   (* check and set outputs *)
     IF #X < #trigger_Low THEN
         #LOW := TRUE;
         #Status := 111;
         IF #Alarm_low THEN
             #Alarm := TRUE;
             #Status := 1;
         END_IF;
     ELSIF #X < #T_1 THEN
         #Q1 := TRUE;
     ELSIF #X < #T_2 THEN
         #Q2 := TRUE;
     ELSIF #X < #T_3 THEN
         #Q3 := TRUE;
     ELSIF #X < #T_4 THEN
         #Q4 := TRUE;
     ELSIF #X < #T_5 THEN
         #Q5 := TRUE;
     ELSIF #X < #trigger_High THEN
         #Q6 := TRUE;
     ELSE
         #HIGH := TRUE;
         #Status := 112;
         IF #Alarm_high THEN
             #Alarm := TRUE;
             #Status := 2;
         END_IF;
     END_IF;

   (* revision history
   hm  22. feb 2007  rev 1.0
     original version

   hm  2. dec 2007   rev 1.1
     chaged code for better performance

   hm  6. jan 2008   rev 1.2
     further performance improvement

   *)
END_FUNCTION_BLOCK

FUNCTION_BLOCK "CALIBRATE"   // FB124, SCL
TITLE = CALIBRATE
{ S7_Optimized_Access := 'FALSE' }
AUTHOR : hugo
FAMILY : MEASURE
NAME : CALIBR
VERSION : 1.3
// Calibrate allows for offset and scale calibration of an analog input.
// offset is calibrated to a stored reference Y_offset while CO is true.
// after the offset is calibrated, scale can be calibrated to a reference value Y_scale while CS is true.
   VAR_INPUT
      X : Real;
      CO : Bool;
      CS : Bool;
      Y_Offset : Real;
      Y_Scale : Real;
   END_VAR
   VAR_OUTPUT
      Y : Real;
   END_VAR
   VAR
      offset : Real;
      Scale : Real := 1.0e+0;
   END_VAR
BEGIN


   (* check for calibration *)
   IF #CO THEN
       #offset := #Y_Offset - #X;
   ELSIF #CS THEN
       #Scale := #Y_Scale / (#X + #offset);
   END_IF;
   (* calculate output *)
   #Y := (#X + #offset) * #Scale;


   (* revision history
   hm 22.2.2007        rev 1.2
       changed VAR RETAIN PERSISTENT to VAR RETAIN for better compatibility
       wago lon contollers do not support persisitent

   hm  11. mar. 2009   rev 1.3
       changed real constants to use dot syntax

   *)
END_FUNCTION_BLOCK

FUNCTION_BLOCK "CYCLE_TIME"   // FB125, SCL
TITLE = CYCLE_TIME
{ S7_Optimized_Access := 'FALSE' }
AUTHOR : hugo
FAMILY : MEASURE
NAME : CYCLE
VERSION : 1.2
// this function block measures the cycle time and displays the last, min and max cycle time of the current task.
// the resolution is 1ms.
// the cycles output is a dword counter which counts the cycles.
// a rst pulse on the input will reset all data.
// 
// uses: T_PLC_MS [FC64]
//       STIME [FB64],IDB_STIME [DB64]
   VAR_INPUT
      rst : Bool;
   END_VAR
   VAR_OUTPUT
      ct_min : Time;
      ct_max : Time;
      ct_last : Time;
      systime : Time;
      sysdays : Int;
      cycles : DWord;
   END_VAR
   VAR
      last_cycle : Time;
      tx : Time;
      init : Bool;
   END_VAR
   VAR_TEMP
      TOP_SI : Struct
         EV_CLASS : Byte;
         EV_NUM : Byte;
         PRIORITY : Byte;
         NUM : Byte;
         TYP2_3 : Byte;
         TYP1 : Byte;
         ZI1 : Word;
         ZI2_3 : DWord;
      END_STRUCT;
      START_UP_SI : Struct
         EV_CLASS : Byte;
         EV_NUM : Byte;
         PRIORITY : Byte;
         NUM : Byte;
         TYP2_3 : Byte;
         TYP1 : Byte;
         ZI1 : Word;
         ZI2_3 : DWord;
      END_STRUCT;
      ERR : Int;
   END_VAR
BEGIN


   (* read actual startup info *)
   (* OB1_SCAN_1  BYTE  -  B#16#01: Abschluss des Neustarts (Warmstarts)
                        -  B#16#02: Abschluss des Wiederanlaufs
                        -  B#16#03: Abschluss des freien Zyklus
                        -  B#16#04: Abschluss des Kaltstarts
                        -  B#16#05: Erster OB 1-Zyklus der neuen Master-CPU nach 
                                    Master-Reserve-Umschaltung und STOP des 
                                    bisherigen Masters *)

     #ERR := RD_SINFO (TOP_SI => #TOP_SI, START_UP_SI => #START_UP_SI);

   (* reset last_time on system startup *)
     IF #TOP_SI.EV_NUM <> 3 THEN 
       #last_cycle := t#0ms;
     END_IF;

     #tx := T_CONV(DWORD_TO_DINT("T_PLC_MS"())) - #last_cycle;

     IF #rst THEN
         #ct_min := t#10h;
         #ct_max := t#0ms;
         #cycles := 0;
     ELSIF #last_cycle > t#0s THEN
         IF #tx < #ct_min THEN #ct_min := #tx;
         ELSIF #tx > #ct_max THEN #ct_max := #tx;
         END_IF;
         #ct_last := #tx;
     ELSIF #ct_min = t#0s THEN
         #ct_min := t#0s - t#1ms;
     END_IF;
     IF #init THEN
         #systime := #systime + #tx;
             IF #systime >= t#1d THEN
                 #systime := #systime - t#1d;
                 #sysdays := #sysdays + 1;
             END_IF;
     END_IF;
     #init := TRUE;
     #last_cycle := #last_cycle + #tx;
     #cycles := DINT_TO_DWORD(DWORD_TO_DINT(#cycles) + 1);

   (*    revision history
   hm 12.12.2006        rev 1.1
       added cycles output, a dword cycle counter.
   hm 10.3.2007         rev 1.2
       changed initialization of ct_min to t#10h for compatibility with siemens s7

   *)
END_FUNCTION_BLOCK

FUNCTION_BLOCK "DT_SIMU"   // FB126, SCL
TITLE = DT_SIMU
{ S7_Optimized_Access := 'FALSE' }
AUTHOR : hugo
FAMILY : MEASURE
NAME : DTSIMU
VERSION : 1.2
// DT_SIMU simulates a real time clock and can be adjusted to different speeds
// it can also be used in simulation to simulate a real time clock.
// the peed of the clock can be increased or decreased to debug timers.
// with the input start a start date-time can be specified.
// 
// uses: AD_DT_TM [FC1]
//       T_PLC_MS [FC64]
//       STIME [FB64],IDB_STIME [DB64]
   VAR_INPUT
      START : Date_And_Time;
      SPEED : Real := 1.0e+0;
   END_VAR
   VAR_OUTPUT
      DTS : Date_And_Time;
   END_VAR
   VAR
      tc : DWord;
      init : Bool;
      last : DWord;
      tx : DWord;
      td : DWord;
   END_VAR
   VAR_TEMP
      TOP_SI : Struct
         EV_CLASS : Byte;
         EV_NUM : Byte;
         PRIORITY : Byte;
         NUM : Byte;
         TYP2_3 : Byte;
         TYP1 : Byte;
         ZI1 : Word;
         ZI2_3 : DWord;
      END_STRUCT;
      START_UP_SI : Struct
         EV_CLASS : Byte;
         EV_NUM : Byte;
         PRIORITY : Byte;
         NUM : Byte;
         TYP2_3 : Byte;
         TYP1 : Byte;
         ZI1 : Word;
         ZI2_3 : DWord;
      END_STRUCT;
      ERR : Int;
   END_VAR
BEGIN


   (* read actual startup info *)
   (* OB1_SCAN_1  BYTE  -  B#16#01: Abschluss des Neustarts (Warmstarts)
                        -  B#16#02: Abschluss des Wiederanlaufs
                        -  B#16#03: Abschluss des freien Zyklus
                        -  B#16#04: Abschluss des Kaltstarts
                        -  B#16#05: Erster OB 1-Zyklus der neuen Master-CPU nach 
                                    Master-Reserve-Umschaltung und STOP des 
                                    bisherigen Masters *)

   #ERR := RD_SINFO (TOP_SI => #TOP_SI, START_UP_SI => #START_UP_SI);

   (* reset last_time on system startup *)
   IF #TOP_SI.EV_NUM = 1 OR #TOP_SI.EV_NUM = 2 OR #TOP_SI.EV_NUM = 4 THEN 
       #init := FALSE;
   END_IF;

   (* read system timer *)
   #tx := "T_PLC_MS"();
   #tc := DINT_TO_DWORD(REAL_TO_DINT(DINT_TO_REAL((DWORD_TO_DINT(#tx) - DWORD_TO_DINT(#last))) * #SPEED));

   IF NOT #init THEN
       #init := TRUE;
       #DTS := #START;
       #tc := 0;
       #last := #tx;
   ELSIF #SPEED = 0.0 THEN
       #DTS := #DTS T_ADD T_CONV(1);
   ELSIF DWORD_TO_DINT(#tc) >= 1000 THEN
       #td := DINT_TO_DWORD((DWORD_TO_DINT(#tc) / 1000)*1000);
       #DTS := #DTS T_ADD T_CONV(DWORD_TO_DINT(#td));
       #last := DINT_TO_DWORD(DWORD_TO_DINT(#last) + REAL_TO_DINT(DINT_TO_REAL(DWORD_TO_DINT(#td)) / #SPEED));
   END_IF;


   (* revision history
   hm  11. sep. 2008   rev 1.0
       original version

   hm  16. nov 2008    rev 1.1
       added type conversions for compatibility reasons

   hm  8.  mar. 2009   rev 1.2
       added increment by cycle mode

   *)
END_FUNCTION_BLOCK

FUNCTION_BLOCK "METER"   // FB127, SCL
TITLE = METER
{ S7_Optimized_Access := 'FALSE' }
AUTHOR : oscat
FAMILY : MEASURE
NAME : METER
VERSION : 1.4
// METER measures usage of power or similar values the output MX is the sum of the inputs over time.
// MX := sum over time of (I1 * P1 + I2 * P2)/D.
// a simple example is the consumption counter for a 2 stage oil burner where stage 1 is 10KW and stage 2 is 20KW.
// I1 and I2 decide which value is accounted for, I1 = True only counts P1, I2 is True counts P2 
// and I1 and I2 is true counts P1 and P2.
// the meter can be used for all kind of consumption meters. P1 and P2 can change on the fly.
// 
// uses: REAL2 [UDT11]
//       T_PLC_MS [FC64]
//       STIME [FB64],IDB_STIME [DB64]
//       R2_ADD [FC144]
   VAR_INPUT
      M1 : Real;
      M2 : Real;
      I1 : Bool;
      I2 : Bool;
      D : Real := 1.0e+0;
      RST : Bool;
   END_VAR
   VAR_IN_OUT
      MX : Real;
   END_VAR
   VAR
      MR : "REAL2";
      MX1 : Real;
      MX2 : Real;
      tx : DWord;
      last : DWord;
      tc : Real;
      init : Bool;
   END_VAR
   VAR_TEMP
      TOP_SI : Struct
         EV_CLASS : Byte;
         EV_NUM : Byte;
         PRIORITY : Byte;
         NUM : Byte;
         TYP2_3 : Byte;
         TYP1 : Byte;
         ZI1 : Word;
         ZI2_3 : DWord;
      END_STRUCT;
      START_UP_SI : Struct
         EV_CLASS : Byte;
         EV_NUM : Byte;
         PRIORITY : Byte;
         NUM : Byte;
         TYP2_3 : Byte;
         TYP1 : Byte;
         ZI1 : Word;
         ZI2_3 : DWord;
      END_STRUCT;
      ERR : Int;
   END_VAR
BEGIN


   (* read actual startup info *)
   (* OB1_SCAN_1  BYTE  -  B#16#01: Abschluss des Neustarts (Warmstarts)
                        -  B#16#02: Abschluss des Wiederanlaufs
                        -  B#16#03: Abschluss des freien Zyklus
                        -  B#16#04: Abschluss des Kaltstarts
                        -  B#16#05: Erster OB 1-Zyklus der neuen Master-CPU nach 
                                    Master-Reserve-Umschaltung und STOP des 
                                    bisherigen Masters *)

   #ERR := RD_SINFO (TOP_SI => #TOP_SI, START_UP_SI => #START_UP_SI);

   (* reset last_time on system startup *)
   IF #TOP_SI.EV_NUM = 1 OR #TOP_SI.EV_NUM = 2 OR #TOP_SI.EV_NUM = 4 THEN 
       #init := FALSE;
   END_IF;

   (* measure the last cycle time and make sure we onle execute once every millisecond *)
   #tx := "T_PLC_MS"();

   IF NOT #init THEN
       #init := TRUE;
       #last := #tx;
       #MR.RX := #MX;
       #MR.R1 := 0.0;
   ELSIF #tx = #last THEN
       RETURN;
   ELSE
       #tc := DINT_TO_REAL(DWORD_TO_DINT(#tx) - DWORD_TO_DINT(#last)) * 0.001;
   END_IF;
   #last := #tx;

   (* reset *)
   IF #RST THEN
       #MR.R1 := 0.0;
       #MR.RX := 0.0;
   ELSE
       (* current consumption measurement *)
       IF #I1 THEN #MX1 := #M1; ELSE #MX1 := 0.0; END_IF;
       IF #I2 THEN #MX2 := #M2; ELSE #MX2 := 0.0; END_IF;
       (* add up the current values in a double real *)
       #MR := "R2_ADD"(X:=#MR,Y:=(SEL(G:=#I1,IN0:=0.0,IN1:=#MX1) + SEL(G:=#I2,IN0:=0.0,IN1:=#MX2)) / #D * #tc);
       (* set the current output value *)
       #MX := #MR.RX;
   END_IF;


   (* revision history

   hm  16. sep.2007        rev 1.0
       original version

   hm  7. feb 2008     rev 1.1
       use new version of ft_int to avoid a counting stop at high values
       deleted unnecessary limits

   hm  24. mar. 2008   rev 1.2
       use data_type real2 to extend accuracy to 15 digits total
       do not use ft_int which adds unnecessary overhead

   hm  8. feb. 2009    rev 1.3
       changed mx to be I/O
       make sure calculation works for cycle times < 1 ms

   hm  8. mar. 2009    rev 1.4
       last was not updated
       code improvements

   *)
END_FUNCTION_BLOCK

FUNCTION_BLOCK "METER_STAT"   // FB128, SCL
TITLE = METER_STAT
{ S7_Optimized_Access := 'FALSE' }
AUTHOR : oscat
FAMILY : MEASURE
NAME : METER_ST
VERSION : 1.3
// METER_STAT runs statistics of a metered value, it calculates the current week, day, month and year consumption and stores the corresponding last day, week, month and year value.
// 
// uses: YEAR_OF_DATE [FC219]
//       MONTH_OF_DATE [FC202]
//       DAY_OF_YEAR [FC180]
//       YEAR_BEGIN [FC217]
//       YEAR_OF_DATE [FC219]
//       LEAP_OF_DATE [FC193] 
//       LEAP_YEAR [FC194]
//       DAY_OF_WEEK [FC179]
   VAR_INPUT
      IN : Real;
      _DI : Date;
      RST : Bool;
   END_VAR
   VAR_IN_OUT
      Last_Day : Real;
      Current_Day : Real;
      Last_Week : Real;
      Current_Week : Real;
      Last_Month : Real;
      Current_Month : Real;
      Last_Year : Real;
      Current_Year : Real;
   END_VAR
   VAR
      Year_Start : Real;
      Month_Start : Real;
      Week_Start : Real;
      Day_Start : Real;
      last_run : Date;
   END_VAR
BEGIN


   IF #RST THEN
       #Last_Day := 0.0;
       #Current_Day := 0.0;
       #Day_Start := #IN;
       #Last_Week := 0.0;
       #Current_Week := 0.0;
       #Week_Start := #IN;
       #Last_Month := 0.0;
       #Current_Month := 0.0;
       #Month_Start := #IN;
       #Last_Year := 0.0;
       #Current_Year := 0.0;
       #Year_Start := #IN;
   ELSE
       #Current_Day := #IN - #Day_Start;
       #Current_Week := #IN - #Week_Start;
       #Current_Month := #IN - #Month_Start;
       #Current_Year := #IN - #Year_Start;
   END_IF;

   IF "YEAR_OF_DATE"(#_DI) > "YEAR_OF_DATE"(#last_run) THEN
       (* a new year has started *)
       #Last_Year := #Current_Year;
       #Current_Year := 0.0;
       #Year_Start := #IN;
       #Last_Month := #Current_Month;
       #Current_Month := 0.0;
       #Month_Start := #IN;
       #Last_Day := #Current_Day;
       #Current_Day := 0.0;
       #Day_Start := #IN;
   ELSIF "MONTH_OF_DATE"(#_DI) > "MONTH_OF_DATE"(#last_run) THEN
       (* a new month has started, january is alrerady done by year change *)
       #Last_Month := #Current_Month;
       #Current_Month := 0.0;
       #Month_Start := #IN;
       #Last_Day := #Current_Day;
       #Current_Day := 0.0;
       #Day_Start := #IN;
   ELSIF "DAY_OF_YEAR"(#_DI) > "DAY_OF_YEAR"(#last_run) THEN
       (* day has chaged, first day of year and first day of month has already been taken care of *)
       #Last_Day := #Current_Day;
       #Current_Day := 0.0;
       #Day_Start := #IN;
   END_IF;
   IF "DAY_OF_WEEK"(#_DI) < "DAY_OF_WEEK"(#last_run) THEN
       (* a new week has started *)
       #Last_Week := #Current_Week;
       #Current_Week := 0.0;
       #Week_Start := #IN;
   END_IF;
   #last_run := #_DI;


   (* revision history
   hm  16. sep. 2007 rev 1.0
     original version

   hm  7. oct. 2008  rev 1.1
     changed function year_to_year_of_date
     changed function month to month_of_date
     changed function weekday to day_of_week

   hm  11. mar. 2009 rev 1.2
     changed real constants to use dot syntax

   hm  18. jul. 2009 rev 1.3
     changes all outputs to be I/O
   *)
END_FUNCTION_BLOCK

FUNCTION_BLOCK "M_D"   // FB129, SCL
TITLE = M_D
{ S7_Optimized_Access := 'FALSE' }
AUTHOR : hugo
FAMILY : MEASURE
NAME : M_D
VERSION : 1.2
// m_d measures the time between a rising edge on start to a rising edge on stop and returs the last measured value on the output PT.
// a second output ET is starting from 0 at the rising edge of start and is counting up until the rising edge of stop occurs.
// the asynchronous input rst can reset the outputs at any time.
// tmax defines a timeout wich is the maximum measurable time between start and stop, if this time is exceeded the outputs will stay at 0.
// 
// uses: T_PLC_MS [FC64]
//       STIME [FB64],IDB_STIME [DB64]
   VAR_INPUT
      start : Bool;
      stop : Bool;
      tmax : Time := T#10D;
      rst : Bool;
   END_VAR
   VAR_OUTPUT
      PT : Time;
      ET : Time;
      run : Bool;
   END_VAR
   VAR
      edge : Bool;
      T_0 : Time;
      tx : Time;
      startup : Bool;
   END_VAR
   VAR_TEMP
      TOP_SI : Struct
         EV_CLASS : Byte;
         EV_NUM : Byte;
         PRIORITY : Byte;
         NUM : Byte;
         TYP2_3 : Byte;
         TYP1 : Byte;
         ZI1 : Word;
         ZI2_3 : DWord;
      END_STRUCT;
      START_UP_SI : Struct
         EV_CLASS : Byte;
         EV_NUM : Byte;
         PRIORITY : Byte;
         NUM : Byte;
         TYP2_3 : Byte;
         TYP1 : Byte;
         ZI1 : Word;
         ZI2_3 : DWord;
      END_STRUCT;
      ERR : Int;
   END_VAR
BEGIN


   (* read actual startup info *)
   (* OB1_SCAN_1  BYTE  -  B#16#01: Abschluss des Neustarts (Warmstarts)
                        -  B#16#02: Abschluss des Wiederanlaufs
                        -  B#16#03: Abschluss des freien Zyklus
                        -  B#16#04: Abschluss des Kaltstarts
                        -  B#16#05: Erster OB 1-Zyklus der neuen Master-CPU nach 
                                    Master-Reserve-Umschaltung und STOP des 
                                    bisherigen Masters *)

   #ERR := RD_SINFO (TOP_SI => #TOP_SI, START_UP_SI => #START_UP_SI);

   (* reset last_time on system startup *)
   IF #TOP_SI.EV_NUM <> 3 THEN 
       #T_0 := t#0ms;
   END_IF;

   (* check for rst input *)
   IF #rst OR #ET >= #tmax THEN
       #PT := t#0ms;
       #ET := t#0ms;
       #startup := FALSE;
       #run := FALSE;
   END_IF;

   (* avoid timers to start when input is true at startup *)
   IF NOT #startup THEN
       #edge := #start;
       #startup := TRUE;
   END_IF;

   (* read system timer *)
   #tx := T_CONV(DWORD_TO_DINT("T_PLC_MS"()));

   (* detect rising edge on start *)
   IF #start AND NOT #edge AND NOT #stop THEN
       #T_0 := #tx;
       #run := TRUE;
       #PT := t#0s;
   ELSIF #stop AND #run THEN
       #PT := #ET;
       #run := FALSE;
   END_IF;
   #edge := #start;
   IF #run THEN #ET := #tx - #T_0; END_IF;


   (* revision history
   hm      2.5.2007    rev 1.0
       original version

   hm        16.9.2007   rev 1.1
       changes time() to T_plc_ms() for compatibility reasons

   hm  27. feb 2009    rev 1.2
       deleted unnecessary init with 0
   *)
END_FUNCTION_BLOCK

FUNCTION_BLOCK "M_T"   // FB130, SCL
TITLE = M_T
{ S7_Optimized_Access := 'FALSE' }
AUTHOR : hugo
FAMILY : MEASURE
NAME : M_T
VERSION : 1.4
// m_t measures the with of a high pulse and returs the last measured pulse width on output PT.
// a second output ET is starting from 0 at the rising edge and counting up until the falling edge occurs and resetts et to 0.
// the asynchrtonous input rst can reset the outputs at any time.
// tmax defines a maximum measurable time, if this value is exceeded the outputs will be reset to 0.
// 
// uses: T_PLC_MS [FC64]
//       STIME [FB64],IDB_STIME [DB64]
   VAR_INPUT
      IN : Bool;
      TMAX : Time := T#10D;
      RST : Bool;
   END_VAR
   VAR_OUTPUT
      PT : Time;
      ET : Time;
   END_VAR
   VAR
      edge : Bool;
      start : Time;
      tx : Time;
   END_VAR
BEGIN


   #tx := T_CONV(DWORD_TO_DINT("T_PLC_MS"()));

   IF #RST OR #ET >= #TMAX THEN
       #PT := t#0s; 
       #ET := t#0s;
   ELSIF #IN THEN
       IF NOT #edge THEN #start := #tx; END_IF;
       #ET := #tx - #start;
   ELSE
       #PT := #ET;
   END_IF;
   #edge := #IN;


   (* revision history
   hm  4. aug. 2006    rev 1.0
       original version

   hm  2. may. 2007    rev 1.1
       added init variable to avoid unreasonable measurement if falling edge occurs first.
       added et (elapsed time) output to count from 0 at rising edge until a falling edge resets et to 0.
       added reset input.

   hm  16. sep. 2007   rev 1.2
       changes time() to T_plc_ms() for compatibility reasons

   hm  17. dec. 2008   rev 1.3
       code optimized

   hm  10. mar. 2009   rev 1.4
       removed nested comments
       removed double assignments

   *)
END_FUNCTION_BLOCK

FUNCTION_BLOCK "M_TX"   // FB131, SCL
TITLE = M_TX
{ S7_Optimized_Access := 'FALSE' }
AUTHOR : oscat
FAMILY : MEASURE
NAME : M_TX
VERSION : 1.4
// this measures the timing of a signal
// TH is the high pulse width
// TL is the low pulse width
// DC is the duty cycle
// F is the frequency
// ET will start at 0 with a rising edge and count up till the next rising edge starts from 0 again. 
// the acuracy depends on the cycle time of the sps and is limited to 1ms resolution.
// an asynchronous reset can reset all outputs to 0 at any time.
// the input tmax can configure a timeout for ET where the function block will outomatically reset itself.
// tmx is predefined to 10 days.
// 
// uses: T_PLC_MS [FC64]
//       STIME [FB64],IDB_STIME [DB64]
   VAR_INPUT
      in : Bool;
      tmax : Time := T#10D;
      rst : Bool;
   END_VAR
   VAR_OUTPUT
      TH : Time;
      TL : Time;
      DC : Real;
      F : Real;
      ET : Time;
   END_VAR
   VAR
      edge : Bool;
      start : Time;
      stop : Time;
      tx : Time;
      rise : Bool;
      fall : Bool;
      startup : Bool;
   END_VAR
BEGIN


   (* check FOR rst input *)
   IF #rst OR (#ET >= #tmax) THEN
       #rise := FALSE;
       #fall := FALSE;
       #startup := FALSE;
       #TH := t#0ms;
       #TL := t#0ms;
       #DC := 0.0;
       #F := 0.0;
       #ET := t#0s;
   END_IF;

   (* avoid timers to start when input is true at startup *)
   IF NOT #startup THEN
       #edge := #in;
       #startup := TRUE;
   END_IF;

   (* read system timer *)
   #tx := T_CONV(DWORD_TO_DINT("T_PLC_MS"()));

   (* edge trigger rising and falling edge *)
   IF #in XOR #edge THEN
       #edge := #in;
       (* rising edge starts measurement *)
       IF #in THEN
           #start := #tx;
           #rise := TRUE;
           IF #fall THEN #TL := #start - #stop; END_IF;
           IF #TH > t#0ms AND #TL > t#0ms THEN
               #DC := DINT_TO_REAL(T_CONV(#TH)) / DINT_TO_REAL(T_CONV(#TH+#TL));
               #F := 1000.0 / DINT_TO_REAL(T_CONV(#TH + #TL));
           END_IF;
       (* falling edge starts second cycle measurement *)
       ELSE
           #stop := #tx;
           #fall := TRUE;
           IF #rise THEN #TH := #stop - #start; END_IF;
           IF #TH > t#0ms AND #TL > t#0ms THEN
               #DC := DINT_TO_REAL(T_CONV(#TH)) /  DINT_TO_REAL(T_CONV(#TH+#TL));
               #F := 1000.0 / DINT_TO_REAL(T_CONV(#TH + #TL));
           END_IF;
       END_IF;
   END_IF;
   IF #rise THEN #ET := #tx - #start; END_IF;


   (* revision history
   hm  4. aug. 2006    rev 1.0
       original version

   hm  2. mai. 2007    rev 1.1
       made sure that no undefined values would be measured at startup conditions
       added output et
       added rst input
       added tmax input

   hm  16. sep. 2007   rev 1.2
       changes time() to T_plc_ms() for compatibility reasons

   hm  27. feb. 2009   rev 1.3
       deleted unnecessary init with 0

   hm  11. mar. 2009   rev 1.4
       changed real constants to use dot syntax

   *)
END_FUNCTION_BLOCK

FUNCTION_BLOCK "ONTIME"   // FB132, SCL
TITLE = ONTIME
{ S7_Optimized_Access := 'FALSE' }
AUTHOR : oscat
FAMILY : MEASURE
NAME : ONTIME
VERSION : 2.5
// ONTIME measures the ontime of a signal in seconds.
// the output SECONDS is of type DWORD which results in a total measurement range of 1 second up to 136 years.
// internally ontime works with a resolution of milliseconds
// 
// uses: T_PLC_MS [FC64]
//       STIME [FB64],IDB_STIME [DB64]
   VAR_INPUT
      IN : Bool;
      RST : Bool;
   END_VAR
   VAR_IN_OUT
      SECONDS : DInt;
      CYCLES : DInt;
   END_VAR
   VAR
      tx : DWord;
      last : DWord;
      edge : Bool;
      init : Bool;
      ms : DWord;
   END_VAR
   VAR_TEMP
      TOP_SI : Struct
         EV_CLASS : Byte;
         EV_NUM : Byte;
         PRIORITY : Byte;
         NUM : Byte;
         TYP2_3 : Byte;
         TYP1 : Byte;
         ZI1 : Word;
         ZI2_3 : DWord;
      END_STRUCT;
      START_UP_SI : Struct
         EV_CLASS : Byte;
         EV_NUM : Byte;
         PRIORITY : Byte;
         NUM : Byte;
         TYP2_3 : Byte;
         TYP1 : Byte;
         ZI1 : Word;
         ZI2_3 : DWord;
      END_STRUCT;
      ERR : Int;
   END_VAR
BEGIN


     (* read actual startup info *)
     (* OB1_SCAN_1  BYTE  -  B#16#01: Abschluss des Neustarts (Warmstarts)
                          -  B#16#02: Abschluss des Wiederanlaufs
                          -  B#16#03: Abschluss des freien Zyklus
                          -  B#16#04: Abschluss des Kaltstarts
                          -  B#16#05: Erster OB 1-Zyklus der neuen Master-CPU nach 
                                      Master-Reserve-Umschaltung und STOP des 
                                      bisherigen Masters *)

     #ERR := RD_SINFO (TOP_SI => #TOP_SI, START_UP_SI => #START_UP_SI);

     (* read system time *)
     #tx := "T_PLC_MS"();

     (* reset last_time on system startup *)
     IF #TOP_SI.EV_NUM = 1 OR #TOP_SI.EV_NUM = 2 OR #TOP_SI.EV_NUM = 4 THEN 
         #init := FALSE;
     END_IF;

     (* make sure the first cycle works correctly *)
     IF NOT #init THEN
       #init := TRUE;
       #last := #tx;
       #ms := 0;
     END_IF;
     IF #RST THEN
       #SECONDS := 0;
       #CYCLES := 0;
       #last := #tx;
       #ms := 0;
     ELSIF #IN THEN
       (* add the current milliseconds *)
       #ms := DINT_TO_DWORD((DWORD_TO_DINT(#tx) - DWORD_TO_DINT(#last)) + DWORD_TO_DINT(#ms));
       IF DWORD_TO_DINT(#ms) >= 1000 THEN
         #SECONDS := #SECONDS + 1;
         #ms := DINT_TO_DWORD(DWORD_TO_DINT(#ms) - 1000);
       END_IF;
       #CYCLES := #CYCLES + BOOL_TO_DINT(NOT #edge);
     END_IF;
     #last := #tx;
     #edge := #IN;


   (* revision history
   hm 22.2.2007    rev 1.1
     changed VAR RETAIN PERSISTENT to VAR RETAIN for better compatibility
     wago lon contollers do not support persisitent

   hm 2.8.2007   rev 1.2
     adding time up in a real number will automatically lead to the point where 
     small time scales like the cycle time will be below the resolution of real and therefore
     ontime would not increase in small steps as necessary
     the time is now measured internally in two  dwords and be converted to real only for
     output purposes.
     deleted the variable power because it was unnecessary

   hm  16.9.2007   rev 1.3
     changes time() to T_plc_ms() for compatibility reasons

   hm  2. dec. 2007  rev 1.4
     chaged code for better performance

   hm  16. mar. 2008 rev 1.5
     added type conversions to avoid warnings under codesys 3.0

   hm  21. oct. 2008 rev 2.0
     changed module for much better performance and allow for external result storage

   hm  10. nov. 2008 rev 2.1
     increased internal resolution to milliseconds

   hm  16. nov. 2008 rev 2.2
     changed typecast to avoid warnings

   hm  17. dec. 2008 rev 2.3
     fixed an error when in would be true for more then 49 days

   hm  17. jan 2011  rev 2.4
     init will not clear seconds and cycles, only rst clears these values  

   hm  18. mar. 2011 rev 2.5
     reset was not working

   *)
END_FUNCTION_BLOCK

FUNCTION_BLOCK "TC_MS"   // FB133, SCL
TITLE = TC_MS
{ S7_Optimized_Access := 'FALSE' }
AUTHOR : hugo
FAMILY : MEASURE
NAME : TC_MS
VERSION : 1.0
// TC_MS delivers the time it was last called on the output TC in Milliseconds.
// 
// uses: T_PLC_MS [FC64]
//       STIME [FB64],IDB_STIME [DB64]
   VAR_OUTPUT
      TC : DWord;
   END_VAR
   VAR
      init : Bool;
      tx : DWord;
      last : DWord;
   END_VAR
   VAR_TEMP
      TOP_SI : Struct
         EV_CLASS : Byte;
         EV_NUM : Byte;
         PRIORITY : Byte;
         NUM : Byte;
         TYP2_3 : Byte;
         TYP1 : Byte;
         ZI1 : Word;
         ZI2_3 : DWord;
      END_STRUCT;
      START_UP_SI : Struct
         EV_CLASS : Byte;
         EV_NUM : Byte;
         PRIORITY : Byte;
         NUM : Byte;
         TYP2_3 : Byte;
         TYP1 : Byte;
         ZI1 : Word;
         ZI2_3 : DWord;
      END_STRUCT;
      ERR : Int;
   END_VAR
BEGIN


   (* read actual startup info *)
   (* OB1_SCAN_1  BYTE  -  B#16#01: Abschluss des Neustarts (Warmstarts)
                        -  B#16#02: Abschluss des Wiederanlaufs
                        -  B#16#03: Abschluss des freien Zyklus
                        -  B#16#04: Abschluss des Kaltstarts
                        -  B#16#05: Erster OB 1-Zyklus der neuen Master-CPU nach 
                                    Master-Reserve-Umschaltung und STOP des 
                                    bisherigen Masters *)

   #ERR := RD_SINFO (TOP_SI => #TOP_SI, START_UP_SI => #START_UP_SI);

   (* reset last_time on system startup *)
   IF #TOP_SI.EV_NUM = 1 OR #TOP_SI.EV_NUM = 2 OR #TOP_SI.EV_NUM = 4 THEN 
       #last := 0;
       #init := FALSE;
   END_IF;

   (* read system timer *)
   #tx := "T_PLC_MS"();

   IF NOT #init THEN
       #init := TRUE;
       #TC := 0;
   ELSE
       #TC := DINT_TO_DWORD(DWORD_TO_DINT(#tx) - DWORD_TO_DINT(#last));
   END_IF;
   #last := #tx;

   (* revision history
   hm      13. mar. 2008   rev 1.0
       original version

   *)
END_FUNCTION_BLOCK

FUNCTION_BLOCK "TC_S"   // FB134, SCL
TITLE = TC_S
{ S7_Optimized_Access := 'FALSE' }
AUTHOR : hugo
FAMILY : MEASURE
NAME : TC_S
VERSION : 1.2
// TC_S delivers the time it was last called on the output TC in seconds.
// 
// uses: T_PLC_US [FC65]
//       STIME [FB64],IDB_STIME [DB64]
   VAR_OUTPUT
      TC : Real;
   END_VAR
   VAR
      init : Bool;
      tx : DWord;
      last : DWord;
   END_VAR
   VAR_TEMP
      TOP_SI : Struct
         EV_CLASS : Byte;
         EV_NUM : Byte;
         PRIORITY : Byte;
         NUM : Byte;
         TYP2_3 : Byte;
         TYP1 : Byte;
         ZI1 : Word;
         ZI2_3 : DWord;
      END_STRUCT;
      START_UP_SI : Struct
         EV_CLASS : Byte;
         EV_NUM : Byte;
         PRIORITY : Byte;
         NUM : Byte;
         TYP2_3 : Byte;
         TYP1 : Byte;
         ZI1 : Word;
         ZI2_3 : DWord;
      END_STRUCT;
      ERR : Int;
   END_VAR
BEGIN


   (* read actual startup info *)
   (* OB1_SCAN_1  BYTE  -  B#16#01: Abschluss des Neustarts (Warmstarts)
                        -  B#16#02: Abschluss des Wiederanlaufs
                        -  B#16#03: Abschluss des freien Zyklus
                        -  B#16#04: Abschluss des Kaltstarts
                        -  B#16#05: Erster OB 1-Zyklus der neuen Master-CPU nach 
                                    Master-Reserve-Umschaltung und STOP des 
                                    bisherigen Masters *)

     #ERR := RD_SINFO (TOP_SI => #TOP_SI, START_UP_SI => #START_UP_SI);

   (* reset last_time on system startup *)
   IF #TOP_SI.EV_NUM = 1 OR #TOP_SI.EV_NUM = 2 OR #TOP_SI.EV_NUM = 4 THEN 
       #last := 0;
       #init := FALSE;
   END_IF;

   (* read system timer *)
   #tx := "T_PLC_US"();

   IF NOT #init THEN
       #init := TRUE;
       #TC := 0.0;
   ELSE
       #TC := (DINT_TO_REAL(DWORD_TO_DINT(#tx)) - DINT_TO_REAL(DWORD_TO_DINT(#last)))*1.0E-6;
   END_IF;
   #last := #tx;


   (* revision history
   hm  13. mar. 2008   rev 1.0
       original version

   hm  16. mar 2008    rev 1.1
       added type conversion to avoid warnings under codesys 3.0

   hm  11. mar. 2009   rev 1.2
       changed real constants to use dot syntax

   *)
END_FUNCTION_BLOCK

FUNCTION_BLOCK "TC_US"   // FB135, SCL
TITLE = TC_US
{ S7_Optimized_Access := 'FALSE' }
AUTHOR : hugo
FAMILY : MEASURE
NAME : TC_US
VERSION : 1.0
// TC_US delivers the time it was last called on the output TC in Microseconds.
// 
// uses: T_PLC_US [FC65]
//       STIME [FB64],IDB_STIME [DB64]
   VAR_OUTPUT
      TC : DWord;
   END_VAR
   VAR
      init : Bool;
      tx : DWord;
      last : DWord;
   END_VAR
   VAR_TEMP
      TOP_SI : Struct
         EV_CLASS : Byte;
         EV_NUM : Byte;
         PRIORITY : Byte;
         NUM : Byte;
         TYP2_3 : Byte;
         TYP1 : Byte;
         ZI1 : Word;
         ZI2_3 : DWord;
      END_STRUCT;
      START_UP_SI : Struct
         EV_CLASS : Byte;
         EV_NUM : Byte;
         PRIORITY : Byte;
         NUM : Byte;
         TYP2_3 : Byte;
         TYP1 : Byte;
         ZI1 : Word;
         ZI2_3 : DWord;
      END_STRUCT;
      ERR : Int;
   END_VAR
BEGIN


   (* read actual startup info *)
   (* OB1_SCAN_1  BYTE  -  B#16#01: Abschluss des Neustarts (Warmstarts)
                        -  B#16#02: Abschluss des Wiederanlaufs
                        -  B#16#03: Abschluss des freien Zyklus
                        -  B#16#04: Abschluss des Kaltstarts
                        -  B#16#05: Erster OB 1-Zyklus der neuen Master-CPU nach 
                                    Master-Reserve-Umschaltung und STOP des 
                                    bisherigen Masters *)

   #ERR := RD_SINFO (TOP_SI => #TOP_SI, START_UP_SI => #START_UP_SI);

   (* reset last_time on system startup *)
   IF #TOP_SI.EV_NUM = 1 OR #TOP_SI.EV_NUM = 2 OR #TOP_SI.EV_NUM = 4 THEN 
       #last := 0;
       #init := FALSE;
   END_IF;

   (* read system timer *)
   #tx := "T_PLC_US"();

   IF NOT #init THEN
       #init := TRUE;
       #TC := 0;
   ELSE
       #TC := DINT_TO_DWORD(DWORD_TO_DINT(#tx) - DWORD_TO_DINT(#last));
   END_IF;
   #last := #tx;

   (* revision history
   hm      13. mar. 2008   rev 1.0
       original version

   *)
END_FUNCTION_BLOCK

FUNCTION_BLOCK "INTEGRATE"   // FB237, SCL
TITLE = INTEGRATE
{ S7_Optimized_Access := 'FALSE' }
AUTHOR : hugo
FAMILY : CTRL
NAME : INTEGR
VERSION : 1.0
// integrate is a plain integrator with I/O for out.
// 
// uses: T_PLC_MS [FC64]
//       STIME [FB64],IDB_STIME [DB64]
   VAR_INPUT
      "E" : Bool := TRUE;
      X : Real;
      K : Real := 1.0e+0;
   END_VAR
   VAR_IN_OUT
      Y : Real;
   END_VAR
   VAR
      X_last : Real;
      init : Bool;
      last : DWord;
      tx : DWord;
   END_VAR
   VAR_TEMP
      TOP_SI : Struct
         EV_CLASS : Byte;
         EV_NUM : Byte;
         PRIORITY : Byte;
         NUM : Byte;
         TYP2_3 : Byte;
         TYP1 : Byte;
         ZI1 : Word;
         ZI2_3 : DWord;
      END_STRUCT;
      START_UP_SI : Struct
         EV_CLASS : Byte;
         EV_NUM : Byte;
         PRIORITY : Byte;
         NUM : Byte;
         TYP2_3 : Byte;
         TYP1 : Byte;
         ZI1 : Word;
         ZI2_3 : DWord;
      END_STRUCT;
      ERR : Int;
   END_VAR
BEGIN


   (* read actual startup info *)
   (* OB1_SCAN_1  BYTE  -  B#16#01: Abschluss des Neustarts (Warmstarts)
                        -  B#16#02: Abschluss des Wiederanlaufs
                        -  B#16#03: Abschluss des freien Zyklus
                        -  B#16#04: Abschluss des Kaltstarts
                        -  B#16#05: Erster OB 1-Zyklus der neuen Master-CPU nach 
                                    Master-Reserve-Umschaltung und STOP des 
                                    bisherigen Masters *)

   #ERR := RD_SINFO (TOP_SI => #TOP_SI, START_UP_SI => #START_UP_SI);

   (* reset last_time on system startup *)
   IF #TOP_SI.EV_NUM = 1 OR #TOP_SI.EV_NUM = 2 OR #TOP_SI.EV_NUM = 4 THEN 
       #init := FALSE;
   END_IF;

   (*read system time *)
   #tx := "T_PLC_MS"();

   IF NOT #init THEN
       #init := TRUE;
       #X_last := #X;
   ELSIF #"E" THEN
       #Y := (#X + #X_last) * 0.5E-3 * DINT_TO_REAL(DWORD_TO_DINT(#tx)-DWORD_TO_DINT(#last)) * #K + #Y;
       #X_last := #X;
   END_IF;
   #last := #tx;


   (*
   hm  3. nov. 2008    rev 1.0
   original version

   *)
END_FUNCTION_BLOCK

FUNCTION_BLOCK "FLOW_METER"   // FB253, SCL
TITLE = FLOW_METER
{ S7_Optimized_Access := 'FALSE' }
AUTHOR : hugo
FAMILY : MEASURE
NAME : FLOWMET
VERSION : 1.0
// Flow meter measures flow according to gated time or pulses.
// 
// uses: INTEGRATE (FB237)
//       T_PLC_MS (FC64)
//       STIME (FB64), IDB_STIME (DB64)
//       FLOOR (FC81)
   VAR_INPUT
      VX : Real;
      "E" : Bool;
      RST : Bool;
      PULSE_MODE : Bool;
      UPDATE_TIME : Time := T#1S;
   END_VAR
   VAR_OUTPUT
      F : Real;
   END_VAR
   VAR_IN_OUT
      X : Real;
      Y : DInt;
   END_VAR
   VAR
      tx : Time;
      tl : Time;
      int1 : "INTEGRATE";
      init : Bool;
      e_last : Bool;
      tmp : Int;
      x_last : Real;
      y_last : DInt;
   END_VAR
   VAR_TEMP
      TOP_SI : Struct
         EV_CLASS : Byte;
         EV_NUM : Byte;
         PRIORITY : Byte;
         NUM : Byte;
         TYP2_3 : Byte;
         TYP1 : Byte;
         ZI1 : Word;
         ZI2_3 : DWord;
      END_STRUCT;
      START_UP_SI : Struct
         EV_CLASS : Byte;
         EV_NUM : Byte;
         PRIORITY : Byte;
         NUM : Byte;
         TYP2_3 : Byte;
         TYP1 : Byte;
         ZI1 : Word;
         ZI2_3 : DWord;
      END_STRUCT;
      ERR : Int;
   END_VAR
BEGIN


   (* read actual startup info *)
   (* OB1_SCAN_1  BYTE  -  B#16#01: Abschluss des Neustarts (Warmstarts)
                        -  B#16#02: Abschluss des Wiederanlaufs
                        -  B#16#03: Abschluss des freien Zyklus
                        -  B#16#04: Abschluss des Kaltstarts
                        -  B#16#05: Erster OB 1-Zyklus der neuen Master-CPU nach 
                                    Master-Reserve-Umschaltung und STOP des 
                                    bisherigen Masters *)

   #ERR := RD_SINFO (TOP_SI => #TOP_SI, START_UP_SI => #START_UP_SI);

   IF NOT #init THEN  (* init on power up *)
     #init := TRUE;
     #tl := #tx;
     #x_last := #X;
     #y_last := #Y;
     #int1.K := 2.7777777777777777E-4;
   END_IF;

   (* run integrator *)
   #int1(E := NOT (#RST OR #PULSE_MODE) AND #"E", X := #VX, Y := #X);  (* gated operation *)

   IF #RST THEN   (* reset *)
     #X := 0.0;
     #Y := 0;
     #tl := #tx;
     #x_last := 0.0;
     #y_last := 0;
   ELSIF #"E" AND #PULSE_MODE THEN  (* check for pulse mode *)
     IF NOT #e_last THEN #X := #X + #VX; END_IF;
   END_IF;
   #e_last := #"E";

   (* reduce X to be less than 1 and increase Y respectively *)
   IF #X > 1.0 THEN
     #tmp := "FLOOR"(#X);
     #Y := #Y + INT_TO_DINT(#tmp);
     #X := #X - INT_TO_REAL(#tmp);
   END_IF;

   (* calculate the current flow *)
   #tx := T_CONV(DWORD_TO_DINT("T_PLC_MS"()));

   (* reset last_time on system startup *)
   IF #TOP_SI.EV_NUM = 1 OR #TOP_SI.EV_NUM = 2 OR #TOP_SI.EV_NUM = 4 THEN 
       #tl := #tx;
   END_IF;

   IF #tx - #tl >= #UPDATE_TIME AND #UPDATE_TIME > t#0s THEN
     #F := (DINT_TO_REAL(#Y - #y_last) + #X - #x_last) / DINT_TO_REAL(T_CONV(#tx - #tl)) * 3.6E6;
     #y_last := #Y;
     #x_last := #X;
     #tl := #tx;
   END_IF;



   (* revision history
   hm  23. jan. 2011 rev 1.0
     original version

   *)
END_FUNCTION_BLOCK

FUNCTION "T_PLC_MS" : DWord   // FC64, SCL
TITLE = T_PLC_MS
{ S7_Optimized_Access := 'FALSE' }
AUTHOR : hugo
FAMILY : MEASURE
NAME : T_PLC_MS
VERSION : 1.2
// T_PLC_MS reads the internal PLC timer and return the time, it has the advantage to be able to set a debug mode 
// and speed up the counter to test the plc timer overrun which occurs every 50 days respectively 25 days at siemens S7
// this routine also allows to correct the behavior of s7 where the internal plc counter will not count all 32 bits.
// 
// uses: STIME [FB64],IDB_STIME [DB64]
BEGIN


   "IDB_STIME"(); 
   #T_PLC_MS := "IDB_STIME".tx; 
   (* hier muss die korrektur für step7 stattfinden
   plctime muss den vollen wertebereich von time ausnutzen:
   wenn bei step7 time -24tage bis plus 24 tage ist dann muss der timer auch beim überlauf auf -24tage springen 
   und auf keinen fall auf 0 !!!!
   für siemens muss ein weiterer fb im main eingebunden werden der sicherstellt das alle 32 bits durchgezählt werden.
   es kann nur ein fb sein den er muss sich das oberste (32te) bit merken.
   oder etwa spring s7 bei überlauf auf -24 tage????? dann wäre keine korrektur nötig.
   *)
   IF "debug" THEN
       #T_PLC_MS := DINT_TO_DWORD((DWORD_TO_DINT(SHL(IN:=#T_PLC_MS,N:="N") OR SHL(IN:=DWORD#1,N:="N"))-1) + DWORD_TO_DINT("offset_1"));
   END_IF;


   (* revision history
   hm  14.9.2007   rev 1.0
       original version

   hm  12. nov 2007    rev 1.1
       added temporaray variable tx because some compilers could not handle time() as an argument

   hm  16. nov. 2008   rev 1.2
       initialized constants with 0 for compatibility reasons
   *)
END_FUNCTION

FUNCTION "T_PLC_US" : DWord   // FC65, SCL
TITLE = T_PLC_US
{ S7_Optimized_Access := 'FALSE' }
AUTHOR : hugo
FAMILY : MEASURE
NAME : T_PLC_US
VERSION : 1.2
// T_PLC_US reads the internal PLC timer and return the time, it has the advantage to be able to set a debug mode 
// and speed up the counter to test the plc timer overrun which occurs every 50 days respectively 25 days at siemens S7
// this routine also allows to correct the behavior of s7 where the internal plc counter will not count all 32 bits.
// 
// uses: STIME [FB64],IDB_STIME [DB64]
BEGIN


   "IDB_STIME"(); 
   #T_PLC_US := DINT_TO_DWORD(DWORD_TO_DINT("IDB_STIME".tx) * 1000); 
   (* hier muss die korrektur für step7 stattfinden
   plctime muss den vollen wertebereich von time ausnutzen:
   wenn bei step7 time -24tage bis plus 24 tage ist dann muss der timer auch beim überlauf auf -24tage springen 
   und auf keinen fall auf 0 !!!!
   für siemens muss ein weiterer fb im main eingebunden werden der sicherstellt das alle 32 bits durchgezählt werden.
   es kann nur ein fb sein den er muss sich das oberste (32te) bit merken.
   oder etwa spring s7 bei überlauf auf -24 tage????? dann wäre keine korrektur nötig.
   *)
   IF "debug" THEN
       #T_PLC_US := DINT_TO_DWORD((DWORD_TO_DINT(SHL(IN:=#T_PLC_US,N:="N") OR SHL(IN:=DWORD#1,N:="N"))-1) + DWORD_TO_DINT("offset_1"));
   END_IF;


   (* revision history
   hm  14.9.2007   rev 1.0
       original version

   hm  12. nov 2007    rev 1.1
       added temporaray variable tx because some compilers could not handle time() as an argument

   hm  16. nov. 2008   rev 1.2
       initialized constants with 0 for compatibility reasons

   *)
END_FUNCTION

FUNCTION "FLOOR" : Int   // FC81, SCL
TITLE = FLOOR
{ S7_Optimized_Access := 'FALSE' }
AUTHOR : hugo
FAMILY : MATH
NAME : FLOOR
VERSION : 1.1
// This is a rounding function which returns the biggest possible integer which is less or equal to X.
// floor(3.14) = 3
// floor(-3.14) = 4
   VAR_INPUT
      X : Real;
   END_VAR
BEGIN


   #FLOOR := REAL_TO_INT(#X);
   IF #FLOOR > #X THEN
       #FLOOR := #FLOOR - 1;
   END_IF;

   (* revision history
   hm    7. feb 2007   rev 1.0
     originlal version

   hm    21. mar. 2008 rev 1.1
     replaced trunc with real_to_int for compatibility reasons

   *)
END_FUNCTION

FUNCTION "R2_ADD" : "REAL2"   // FC144, SCL
TITLE = R2_ADD
{ S7_Optimized_Access := 'FALSE' }
AUTHOR : hugo
FAMILY : R2
NAME : ADD
VERSION : 1.0
// R2_add adds a real to a double real which extends the accuracy of a real to twice as many digits
//  
// uses: REAL2 [UDT11]
   VAR_INPUT
      X : "REAL2";
      Y : Real;
   END_VAR
   VAR_TEMP
      temp : Real;
      tR2_ADD : "REAL2";
   END_VAR
BEGIN


   #temp := #X.RX;
   #tR2_ADD.RX := #Y + #X.R1 + #X.RX;
   #tR2_ADD.R1 := #temp - #tR2_ADD.RX + #Y + #X.R1;

   #R2_ADD := #tR2_ADD;

   (* revision history
   hm      20.3.2008   rev 1.0
       original version

   *)
END_FUNCTION

FUNCTION "DAY_OF_WEEK" : Int   // FC179, SCL
TITLE = DAY_OF_WEEK
{ S7_Optimized_Access := 'FALSE' }
AUTHOR : hugo
FAMILY : TIDT
NAME : DWEEK
VERSION : 1.4
// calculates the weekday of a week according to ISO8601   
// monday = 1 ..... sunday = 7
   VAR_INPUT
      IDATE : Date;
   END_VAR
BEGIN


     #DAY_OF_WEEK := DINT_TO_INT((T_CONV(#IDATE)+7308) MOD 7)+1;

   (* 
   weekday := DWORD_TO_INT((DATE_TO_DWORD(idate)/86400+3) MOD 7) + 1;
   *)


   (* revision history
   hm  21.8.06         rev 1.1
       corrected a miscalculation

   hm  23.12.2007      rev 1.2
       correction for step7

   hm  7. apr. 2008    rev 1.3
       deleted unused step7 code

   hm  7. oct. 2008    rev 1.4
       changed name of function from weekday to day_of_week

   *)
END_FUNCTION

FUNCTION "DAY_OF_YEAR" : Int   // FC180, SCL
TITLE = DAY_OF_YEAR
{ S7_Optimized_Access := 'FALSE' }
AUTHOR : hugo
FAMILY : TIDT
NAME : DAYOYEAR
VERSION : 1.4
// calculates the day of the year
// 
// uses: DATE_DINT [FC405]
   VAR_INPUT
      idate : Date;
   END_VAR
BEGIN


   #DAY_OF_YEAR := DINT_TO_INT(("DATE_DINT"(#idate) / 86400) MOD 1461);
   IF #DAY_OF_YEAR > 729 THEN
     IF #DAY_OF_YEAR > 1095 THEN #DAY_OF_YEAR := #DAY_OF_YEAR - 1095; ELSE #DAY_OF_YEAR := #DAY_OF_YEAR - 729; END_IF;
   ELSIF #DAY_OF_YEAR > 364 THEN
     #DAY_OF_YEAR := #DAY_OF_YEAR - 364;
   ELSE
     #DAY_OF_YEAR := #DAY_OF_YEAR + 1;
   END_IF;

   //  day_of_year := DINT_TO_INT((DATE_TO_DINT(idate) - DATE_TO_DINT(year_begin(year_of_date(idate))))) + 1;

   (*
   DAY_OF_YEAR := DWORD_TO_INT((DATE_TO_DWORD(idate) - DATE_TO_DWORD(YEAR_BEGIN(YEAR_OF_DATE(idate)))) / 86400) + 1;
   *)


   (* revivision history
   hm  4. aug. 2007    rev 1.0
     original version

   hm  1. oct. 2007    rev 1.1
     added compatibility to STEP7

   hm  4. jan. 2008    rev 1.2
     changed code for better performance

   hm  7. oct. 2008    rev 1.3
     changed name of function year to year_of_date

   hm  28. jan. 2011 rev 1.4
     improved code
   *)
END_FUNCTION

FUNCTION "LEAP_OF_DATE" : Bool   // FC193, SCL
TITLE = LEAP_OF_DATE
{ S7_Optimized_Access := 'FALSE' }
AUTHOR : hugo
FAMILY : TIDT
NAME : LEAPODAT
VERSION : 1.3
// leap_year is true if the tested year is a leap year  
// 
// uses: DATE_DINT [FC405]
   VAR_INPUT
      idate : Date;
   END_VAR
BEGIN


   #LEAP_OF_DATE := SHL(IN:=DINT_TO_DWORD((("DATE_DINT"(#idate) + 43200) / 31557600)),N:=30) = 16#80000000;


   (* change history

   2.10.2006   rev 1.1
   the function now calls leap_year to accomodate further accuracy.
   the function now works for any year from 1970 to 2100

   8. jan 2008   rev 1.2
     improved code for better performance

   28. jan. 2011 rev 1.3
     improved performance
   *)
END_FUNCTION

FUNCTION "MONTH_OF_DATE" : Int   // FC202, SCL
TITLE = MONTH_OF_DATE
{ S7_Optimized_Access := 'FALSE' }
AUTHOR : hugo
FAMILY : TIDT
NAME : MONTH
VERSION : 1.3
// returns the month of a date  
// 
// uses: DAY_OF_YEAR [FC180]
//       YEAR_BEGIN [FC217] 
//       YEAR_OF_DATE [FC219] 
//       LEAP_OF_DATE [FC193]
//       LEAP_YEAR [FC194]
   VAR_INPUT
      IDATE : Date;
   END_VAR
BEGIN


   #MONTH_OF_DATE := "DAY_OF_YEAR"(#IDATE);
   IF #MONTH_OF_DATE < 32 THEN
       #MONTH_OF_DATE := 1;
   ELSIF "LEAP_OF_DATE"(#IDATE) THEN
       #MONTH_OF_DATE := (#MONTH_OF_DATE * 53 + 1668) / 1623;
   ELSE
       #MONTH_OF_DATE := (#MONTH_OF_DATE * 53 + 1700) / 1620;
   END_IF;


   (* code for rev 1.2
   MONTH_OF_DATE := DAY_OF_YEAR(IDATE);
   IF LEAP_OF_DATE(IDATE) THEN
       CASE MONTH_OF_DATE OF
           1..31   :   MONTH_OF_DATE := 1;
           32..60  :   MONTH_OF_DATE := 2;
           61..91  :   MONTH_OF_DATE := 3;
           92..121 :   MONTH_OF_DATE := 4;
           122..152:   MONTH_OF_DATE := 5;
           153..182:   MONTH_OF_DATE := 6;
           183..213:   MONTH_OF_DATE := 7;
           214..244:   MONTH_OF_DATE := 8;
           245..274:   MONTH_OF_DATE := 9;
           275..305:   MONTH_OF_DATE := 10;
           306..335:   MONTH_OF_DATE := 11;
           336..366:   MONTH_OF_DATE := 12;
       END_CASE;
   ELSE
       CASE MONTH_OF_DATE OF
           1..31   :   MONTH_OF_DATE := 1;
           32..59  :   MONTH_OF_DATE := 2;
           60..90  :   MONTH_OF_DATE := 3;
           91..120 :   MONTH_OF_DATE := 4;
           121..151:   MONTH_OF_DATE := 5;
           152..181:   MONTH_OF_DATE := 6;
           182..212:   MONTH_OF_DATE := 7;
           213..243:   MONTH_OF_DATE := 8;
           244..273:   MONTH_OF_DATE := 9;
           274..304:   MONTH_OF_DATE := 10;
           305..334:   MONTH_OF_DATE := 11;
           335..365:   MONTH_OF_DATE := 12;
       END_CASE;
   END_IF;
   *)


   (* revision history
   hm  1. aug 2006 rev 1.0
       original version    

   hm  1. okt 2007 rev 1.1
       replaced old code (string conversion) with mathematics
       the execution time is now multiple times faster.

   hm  7. oct. 2008    rev 1.2
       changed name of function from month to MONTH_OF_DATE

   hm  27. mar. 2009   rev 1.3
       new improved code

   *)
END_FUNCTION

FUNCTION "YEAR_OF_DATE" : Int   // FC219, SCL
TITLE = YEAR_OF_DATE
{ S7_Optimized_Access := 'FALSE' }
AUTHOR : hugo
FAMILY : TIDT
NAME : YEAR
VERSION : 1.4
// returs the year of a date  
// the function works for dates from 1990 - 2100
   VAR_INPUT
      IDATE : Date;
   END_VAR
BEGIN


   #YEAR_OF_DATE := DINT_TO_INT(((100 * T_CONV(#IDATE)) + 50) / 36525) + 1990;  

   (*
   year := DWORD_TO_INT((DATE_TO_DWORD(idate)+43200) / 31557600 + 1970);
   *)

   (* code used prior to rev 1.1
   year := DWORD_TO_INT((DATE_TO_DWORD(idate)/864+71954300)/36525);
   *)

   (* revision history
   hm  4. aug 2006     rev 1.0
       original version

   hm  1. okt 2007     rev 1.1
       corrected error in algorithm
       adjustment for S7 compatibility

   hm  23.12.2007      rev 1.2
       changed code for better performance

   hm  7. apr. 2008    rev 1.3
       deleted unused step7 code

   hm  7. oct. 2008    rev 1.4
       reneamed function (year) to year_of_date

   *)
END_FUNCTION

FUNCTION "DATE_DINT" : DInt   // FC405, SCL
TITLE = DATE_DINT
{ S7_Optimized_Access := 'FALSE' }
AUTHOR : dalbi
FAMILY : xS7
NAME : D_DINT
VERSION : 1.0
// convert S7 DATE to IEC-DATE
   VAR_INPUT
      D : Date;
   END_VAR
BEGIN


   (* 1.1.1990 00:00:00 = 631152000 *)
   #DATE_DINT := T_CONV(#D) * 86400 + 631152000;
END_FUNCTION

// ===== PLC "Engineering sensor"  Unspecific CPU S7 300 =====
